(* Logix 5000 project; controller PLC_MCC1300_75F1 vendor 1 type 14 code 166 rev 32.11; software revision 32.04; part 47 of 83 *)
(* tags used below, declared in another part *)
   GP_TrackingFiring : GP_TrackingFiring;
   GP_TrackingFiringForConvoy : GP_TrackingFiringForConvoy;
   M30xTrimWheel : MAC_TrimmingWheels[5];
   M30xTrimWheel_HMR : MAC_TrimmingWheels_HMR[5];
   M30xTrimWheel_HMW : MAC_TrimmingWheels_HMW[5];
   TMP_d : DINT;
   TMP_dIndex : DINT;
   xAlwaysOFF : BOOL;
   Z300_BufferPlate : UDT_LINE_BUFFER_PLATE;
   Z301 : MAC_Zone_ML;
(* MainProgram, continued *)

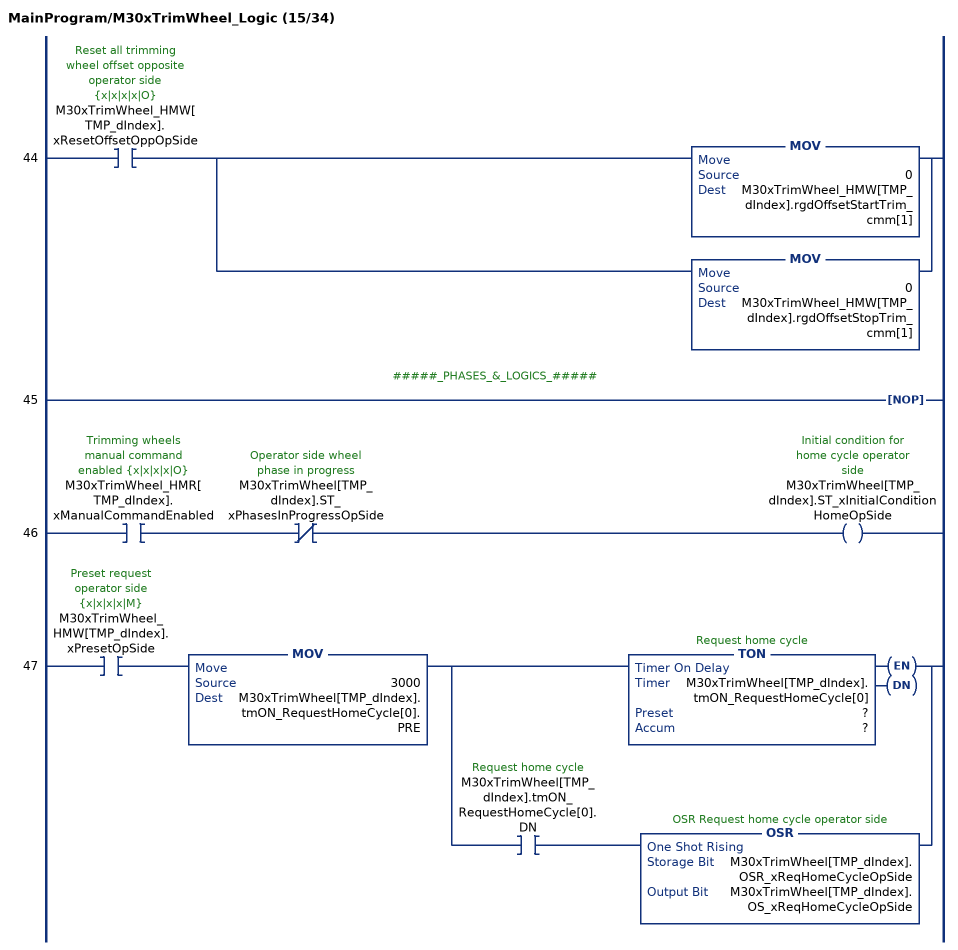
   [picture p701: MainProgram/M30xTrimWheel_Logic rungs 44-47]
   44: XIC(M30xTrimWheel_HMW[TMP_dIndex].xResetOffsetOppOpSide)[MOV(0,M30xTrimWheel_HMW[TMP_dIndex].rgdOffsetStartTrim_cmm[1]) ,MOV(0,M30xTrimWheel_HMW[TMP_dIndex].rgdOffsetStopTrim_cmm[1]) ];
   // #####_PHASES_&_LOGICS_#####
   45: NOP();
   46: XIC(M30xTrimWheel_HMR[TMP_dIndex].xManualCommandEnabled)XIO(M30xTrimWheel[TMP_dIndex].ST_xPhasesInProgressOpSide)OTE(M30xTrimWheel[TMP_dIndex].ST_xInitialConditionHomeOpSide);
   47: XIC(M30xTrimWheel_HMW[TMP_dIndex].xPresetOpSide)MOV(3000,M30xTrimWheel[TMP_dIndex].tmON_RequestHomeCycle[0].PRE)[TON(M30xTrimWheel[TMP_dIndex].tmON_RequestHomeCycle[0],?,?) ,XIC(M30xTrimWheel[TMP_dIndex].tmON_RequestHomeCycle[0].DN) OSR(M30xTrimWheel[TMP_dIndex].OSR_xReqHomeCycleOpSide,M30xTrimWheel[TMP_dIndex].OS_xReqHomeCycleOpSide) ];
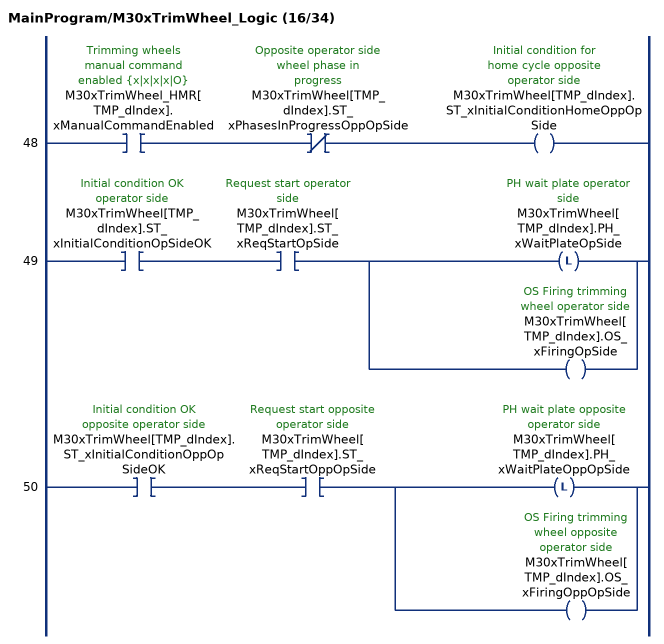
   48: XIC(M30xTrimWheel_HMR[TMP_dIndex].xManualCommandEnabled)XIO(M30xTrimWheel[TMP_dIndex].ST_xPhasesInProgressOppOpSide)OTE(M30xTrimWheel[TMP_dIndex].ST_xInitialConditionHomeOppOpSide);
   49: XIC(M30xTrimWheel[TMP_dIndex].ST_xInitialConditionOpSideOK)XIC(M30xTrimWheel[TMP_dIndex].ST_xReqStartOpSide)[OTL(M30xTrimWheel[TMP_dIndex].PH_xWaitPlateOpSide) ,OTE(M30xTrimWheel[TMP_dIndex].OS_xFiringOpSide) ];
   50: XIC(M30xTrimWheel[TMP_dIndex].ST_xInitialConditionOppOpSideOK)XIC(M30xTrimWheel[TMP_dIndex].ST_xReqStartOppOpSide)[OTL(M30xTrimWheel[TMP_dIndex].PH_xWaitPlateOppOpSide) ,OTE(M30xTrimWheel[TMP_dIndex].OS_xFiringOppOpSide) ];
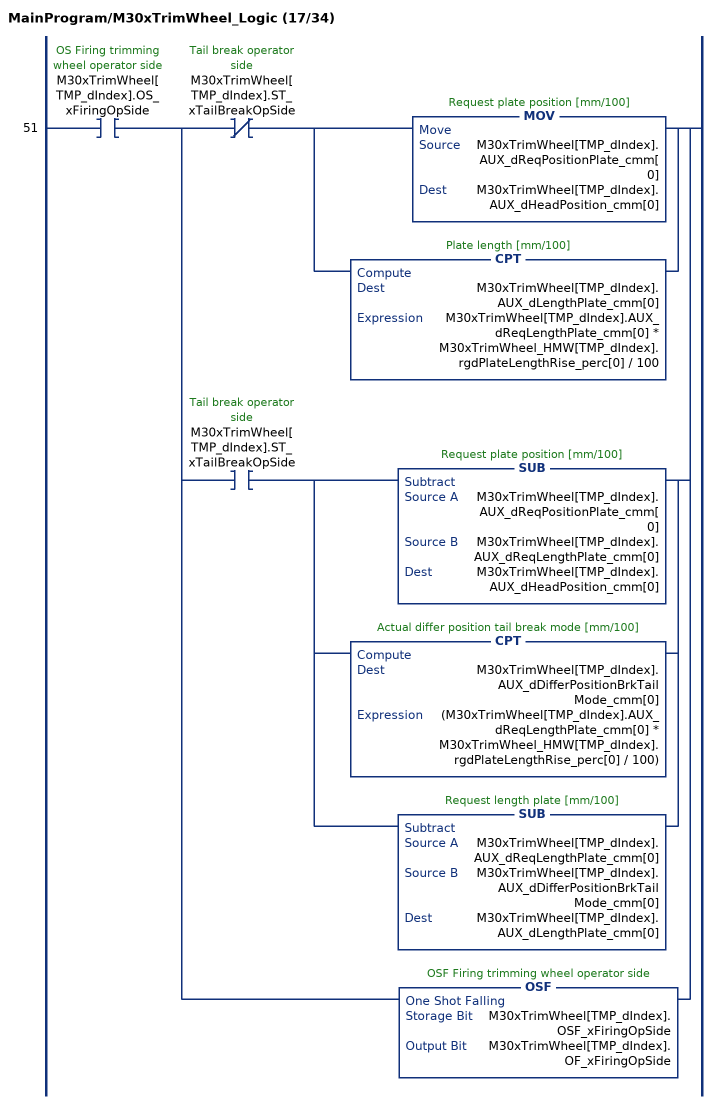
   51: XIC(M30xTrimWheel[TMP_dIndex].OS_xFiringOpSide)[XIO(M30xTrimWheel[TMP_dIndex].ST_xTailBreakOpSide) [MOV(M30xTrimWheel[TMP_dIndex].AUX_dReqPositionPlate_cmm[0],M30xTrimWheel[TMP_dIndex].AUX_dHeadPosition_cmm[0]) ,CPT(M30xTrimWheel[TMP_dIndex].AUX_dLengthPlate_cmm[0],M30xTrimWheel[TMP_dIndex].AUX_dReqLengthPlate_cmm[0] * M30xTrimWheel_HMW[TMP_dIndex].rgdPlateLengthRise_perc[0] / 100) ] ,XIC(M30xTrimWheel[TMP_dIndex].ST_xTailBreakOpSide) [SUB(M30xTrimWheel[TMP_dIndex].AUX_dReqPositionPlate_cmm[0],M30xTrimWheel[TMP_dIndex].AUX_dReqLengthPlate_cmm[0],M30xTrimWheel[TMP_dIndex].AUX_dHeadPosition_cmm[0]) ,CPT(M30xTrimWheel[TMP_dIndex].AUX_dDifferPositionBrkTailMode_cmm[0],(M30xTrimWheel[TMP_dIndex].AUX_dReqLengthPlate_cmm[0] * M30xTrimWheel_HMW[TMP_dIndex].rgdPlateLengthRise_perc[0] / 100)) ,SUB(M30xTrimWheel[TMP_dIndex].AUX_dReqLengthPlate_cmm[0],M30xTrimWheel[TMP_dIndex].AUX_dDifferPositionBrkTailMode_cmm[0],M30xTrimWheel[TMP_dIndex].AUX_dLengthPlate_cmm[0]) ] ,OSF(M30xTrimWheel[TMP_dIndex].OSF_xFiringOpSide,M30xTrimWheel[TMP_dIndex].OF_xFiringOpSide) ];
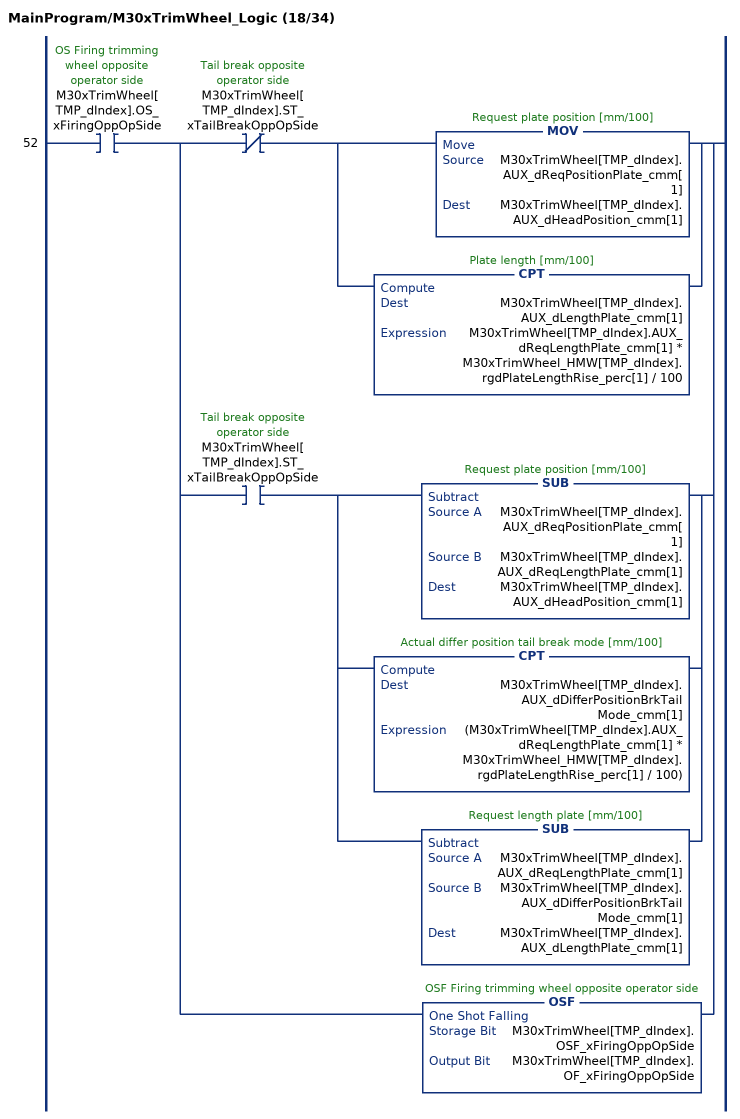
   52: XIC(M30xTrimWheel[TMP_dIndex].OS_xFiringOppOpSide)[XIO(M30xTrimWheel[TMP_dIndex].ST_xTailBreakOppOpSide) [MOV(M30xTrimWheel[TMP_dIndex].AUX_dReqPositionPlate_cmm[1],M30xTrimWheel[TMP_dIndex].AUX_dHeadPosition_cmm[1]) ,CPT(M30xTrimWheel[TMP_dIndex].AUX_dLengthPlate_cmm[1],M30xTrimWheel[TMP_dIndex].AUX_dReqLengthPlate_cmm[1] * M30xTrimWheel_HMW[TMP_dIndex].rgdPlateLengthRise_perc[1] / 100) ] ,XIC(M30xTrimWheel[TMP_dIndex].ST_xTailBreakOppOpSide) [SUB(M30xTrimWheel[TMP_dIndex].AUX_dReqPositionPlate_cmm[1],M30xTrimWheel[TMP_dIndex].AUX_dReqLengthPlate_cmm[1],M30xTrimWheel[TMP_dIndex].AUX_dHeadPosition_cmm[1]) ,CPT(M30xTrimWheel[TMP_dIndex].AUX_dDifferPositionBrkTailMode_cmm[1],(M30xTrimWheel[TMP_dIndex].AUX_dReqLengthPlate_cmm[1] * M30xTrimWheel_HMW[TMP_dIndex].rgdPlateLengthRise_perc[1] / 100)) ,SUB(M30xTrimWheel[TMP_dIndex].AUX_dReqLengthPlate_cmm[1],M30xTrimWheel[TMP_dIndex].AUX_dDifferPositionBrkTailMode_cmm[1],M30xTrimWheel[TMP_dIndex].AUX_dLengthPlate_cmm[1]) ] ,OSF(M30xTrimWheel[TMP_dIndex].OSF_xFiringOppOpSide,M30xTrimWheel[TMP_dIndex].OF_xFiringOppOpSide) ];
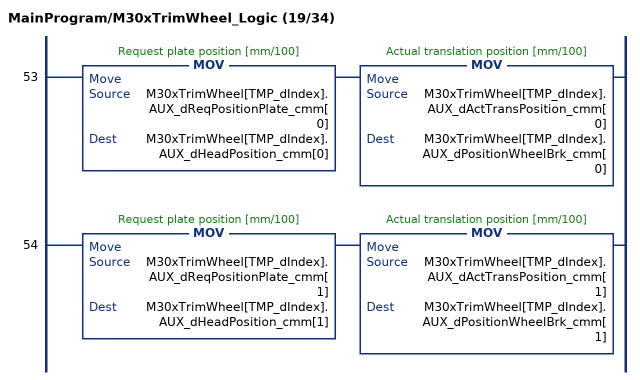
   53: MOV(M30xTrimWheel[TMP_dIndex].AUX_dReqPositionPlate_cmm[0],M30xTrimWheel[TMP_dIndex].AUX_dHeadPosition_cmm[0])MOV(M30xTrimWheel[TMP_dIndex].AUX_dActTransPosition_cmm[0],M30xTrimWheel[TMP_dIndex].AUX_dPositionWheelBrk_cmm[0]);
   54: MOV(M30xTrimWheel[TMP_dIndex].AUX_dReqPositionPlate_cmm[1],M30xTrimWheel[TMP_dIndex].AUX_dHeadPosition_cmm[1])MOV(M30xTrimWheel[TMP_dIndex].AUX_dActTransPosition_cmm[1],M30xTrimWheel[TMP_dIndex].AUX_dPositionWheelBrk_cmm[1]);
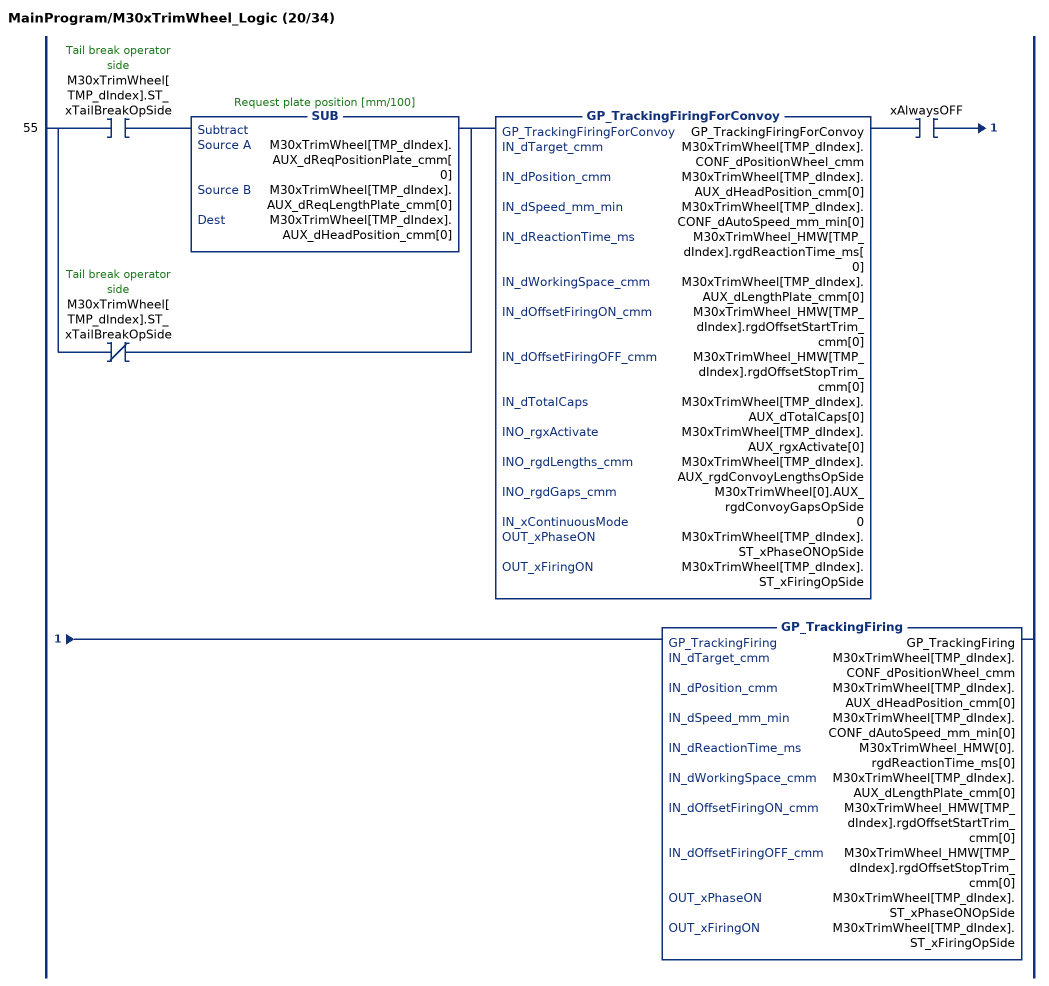
   55: [XIC(M30xTrimWheel[TMP_dIndex].ST_xTailBreakOpSide) SUB(M30xTrimWheel[TMP_dIndex].AUX_dReqPositionPlate_cmm[0],M30xTrimWheel[TMP_dIndex].AUX_dReqLengthPlate_cmm[0],M30xTrimWheel[TMP_dIndex].AUX_dHeadPosition_cmm[0]) ,XIO(M30xTrimWheel[TMP_dIndex].ST_xTailBreakOpSide) ]GP_TrackingFiringForConvoy(GP_TrackingFiringForConvoy,M30xTrimWheel[TMP_dIndex].CONF_dPositionWheel_cmm,M30xTrimWheel[TMP_dIndex].AUX_dHeadPosition_cmm[0],M30xTrimWheel[TMP_dIndex].CONF_dAutoSpeed_mm_min[0],M30xTrimWheel_HMW[TMP_dIndex].rgdReactionTime_ms[0],M30xTrimWheel[TMP_dIndex].AUX_dLengthPlate_cmm[0],M30xTrimWheel_HMW[TMP_dIndex].rgdOffsetStartTrim_cmm[0],M30xTrimWheel_HMW[TMP_dIndex].rgdOffsetStopTrim_cmm[0],M30xTrimWheel[TMP_dIndex].AUX_dTotalCaps[0],M30xTrimWheel[TMP_dIndex].AUX_rgxActivate[0],M30xTrimWheel[TMP_dIndex].AUX_rgdConvoyLengthsOpSide,M30xTrimWheel[0].AUX_rgdConvoyGapsOpSide,0,M30xTrimWheel[TMP_dIndex].ST_xPhaseONOpSide,M30xTrimWheel[TMP_dIndex].ST_xFiringOpSide)XIC(xAlwaysOFF)GP_TrackingFiring(GP_TrackingFiring,M30xTrimWheel[TMP_dIndex].CONF_dPositionWheel_cmm,M30xTrimWheel[TMP_dIndex].AUX_dHeadPosition_cmm[0],M30xTrimWheel[TMP_dIndex].CONF_dAutoSpeed_mm_min[0],M30xTrimWheel_HMW[0].rgdReactionTime_ms[0],M30xTrimWheel[TMP_dIndex].AUX_dLengthPlate_cmm[0],M30xTrimWheel_HMW[TMP_dIndex].rgdOffsetStartTrim_cmm[0],M30xTrimWheel_HMW[TMP_dIndex].rgdOffsetStopTrim_cmm[0],M30xTrimWheel[TMP_dIndex].ST_xPhaseONOpSide,M30xTrimWheel[TMP_dIndex].ST_xFiringOpSide);
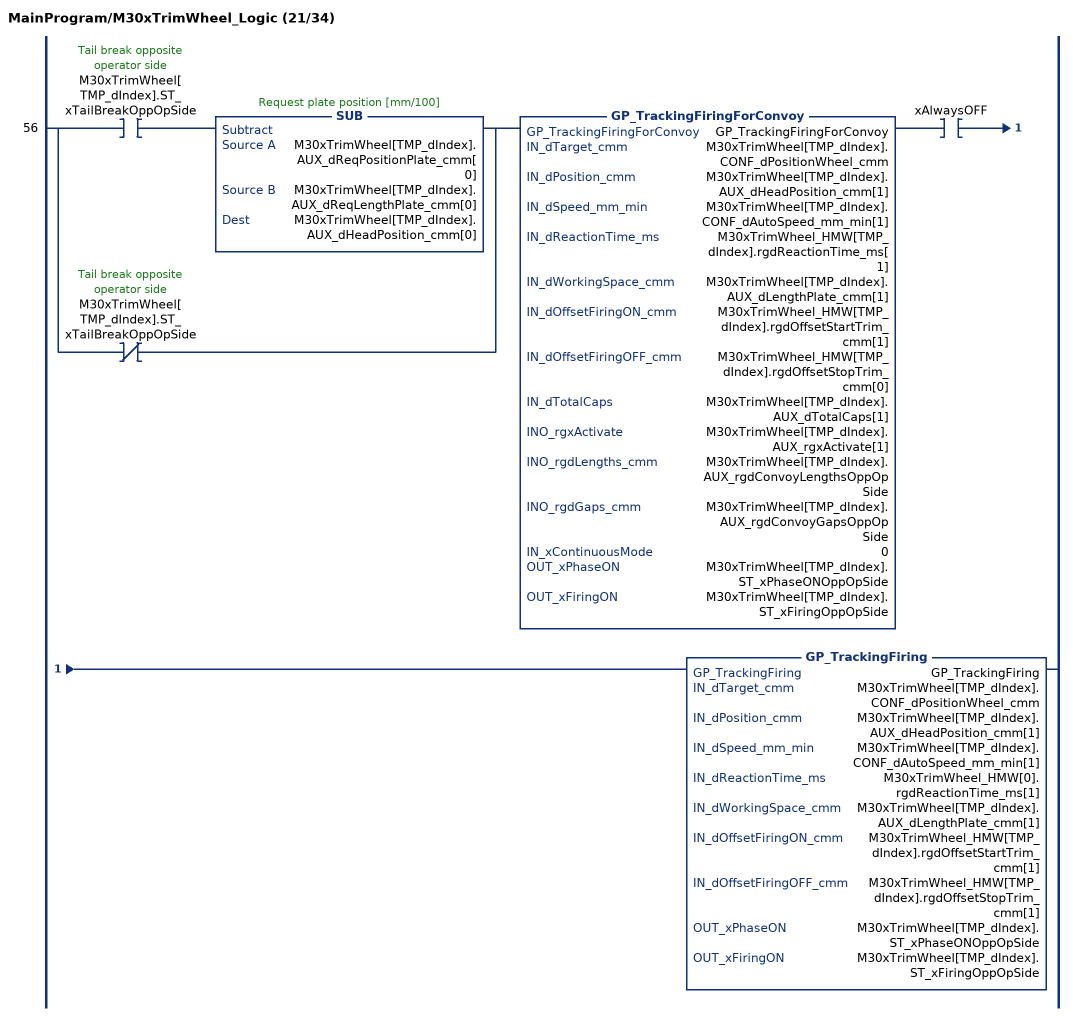
   56: [XIC(M30xTrimWheel[TMP_dIndex].ST_xTailBreakOppOpSide) SUB(M30xTrimWheel[TMP_dIndex].AUX_dReqPositionPlate_cmm[0],M30xTrimWheel[TMP_dIndex].AUX_dReqLengthPlate_cmm[0],M30xTrimWheel[TMP_dIndex].AUX_dHeadPosition_cmm[0]) ,XIO(M30xTrimWheel[TMP_dIndex].ST_xTailBreakOppOpSide) ]GP_TrackingFiringForConvoy(GP_TrackingFiringForConvoy,M30xTrimWheel[TMP_dIndex].CONF_dPositionWheel_cmm,M30xTrimWheel[TMP_dIndex].AUX_dHeadPosition_cmm[1],M30xTrimWheel[TMP_dIndex].CONF_dAutoSpeed_mm_min[1],M30xTrimWheel_HMW[TMP_dIndex].rgdReactionTime_ms[1],M30xTrimWheel[TMP_dIndex].AUX_dLengthPlate_cmm[1],M30xTrimWheel_HMW[TMP_dIndex].rgdOffsetStartTrim_cmm[1],M30xTrimWheel_HMW[TMP_dIndex].rgdOffsetStopTrim_cmm[0],M30xTrimWheel[TMP_dIndex].AUX_dTotalCaps[1],M30xTrimWheel[TMP_dIndex].AUX_rgxActivate[1],M30xTrimWheel[TMP_dIndex].AUX_rgdConvoyLengthsOppOpSide,M30xTrimWheel[TMP_dIndex].AUX_rgdConvoyGapsOppOpSide,0,M30xTrimWheel[TMP_dIndex].ST_xPhaseONOppOpSide,M30xTrimWheel[TMP_dIndex].ST_xFiringOppOpSide)XIC(xAlwaysOFF)GP_TrackingFiring(GP_TrackingFiring,M30xTrimWheel[TMP_dIndex].CONF_dPositionWheel_cmm,M30xTrimWheel[TMP_dIndex].AUX_dHeadPosition_cmm[1],M30xTrimWheel[TMP_dIndex].CONF_dAutoSpeed_mm_min[1],M30xTrimWheel_HMW[0].rgdReactionTime_ms[1],M30xTrimWheel[TMP_dIndex].AUX_dLengthPlate_cmm[1],M30xTrimWheel_HMW[TMP_dIndex].rgdOffsetStartTrim_cmm[1],M30xTrimWheel_HMW[TMP_dIndex].rgdOffsetStopTrim_cmm[1],M30xTrimWheel[TMP_dIndex].ST_xPhaseONOppOpSide,M30xTrimWheel[TMP_dIndex].ST_xFiringOppOpSide);
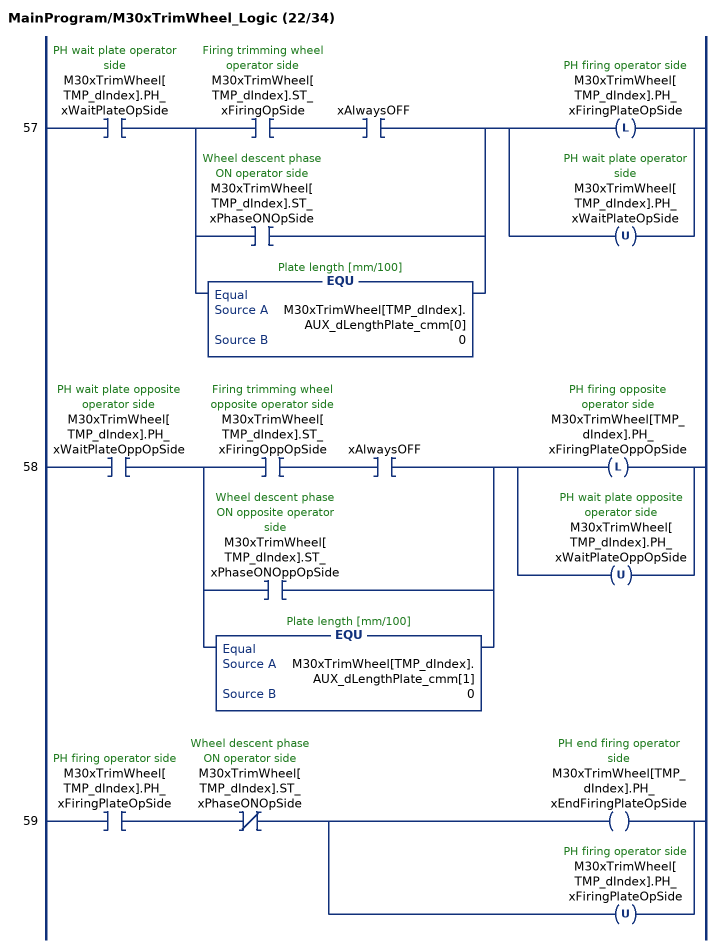
   57: XIC(M30xTrimWheel[TMP_dIndex].PH_xWaitPlateOpSide)[XIC(M30xTrimWheel[TMP_dIndex].ST_xFiringOpSide) XIC(xAlwaysOFF) ,XIC(M30xTrimWheel[TMP_dIndex].ST_xPhaseONOpSide) ,EQU(M30xTrimWheel[TMP_dIndex].AUX_dLengthPlate_cmm[0],0) ][OTL(M30xTrimWheel[TMP_dIndex].PH_xFiringPlateOpSide) ,OTU(M30xTrimWheel[TMP_dIndex].PH_xWaitPlateOpSide) ];
   58: XIC(M30xTrimWheel[TMP_dIndex].PH_xWaitPlateOppOpSide)[XIC(M30xTrimWheel[TMP_dIndex].ST_xFiringOppOpSide) XIC(xAlwaysOFF) ,XIC(M30xTrimWheel[TMP_dIndex].ST_xPhaseONOppOpSide) ,EQU(M30xTrimWheel[TMP_dIndex].AUX_dLengthPlate_cmm[1],0) ][OTL(M30xTrimWheel[TMP_dIndex].PH_xFiringPlateOppOpSide) ,OTU(M30xTrimWheel[TMP_dIndex].PH_xWaitPlateOppOpSide) ];
   59: XIC(M30xTrimWheel[TMP_dIndex].PH_xFiringPlateOpSide)XIO(M30xTrimWheel[TMP_dIndex].ST_xPhaseONOpSide)[OTE(M30xTrimWheel[TMP_dIndex].PH_xEndFiringPlateOpSide) ,OTU(M30xTrimWheel[TMP_dIndex].PH_xFiringPlateOpSide) ];
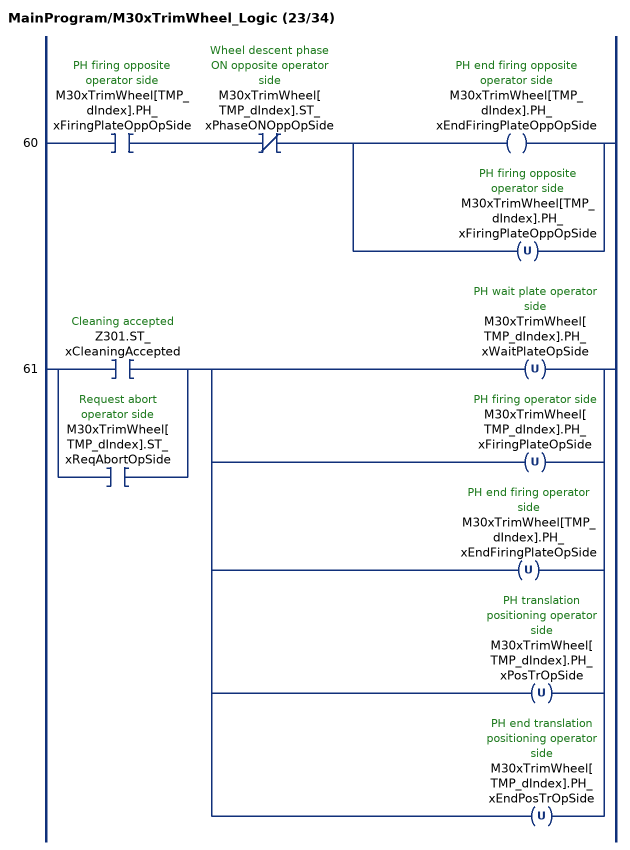
   60: XIC(M30xTrimWheel[TMP_dIndex].PH_xFiringPlateOppOpSide)XIO(M30xTrimWheel[TMP_dIndex].ST_xPhaseONOppOpSide)[OTE(M30xTrimWheel[TMP_dIndex].PH_xEndFiringPlateOppOpSide) ,OTU(M30xTrimWheel[TMP_dIndex].PH_xFiringPlateOppOpSide) ];
   61: [XIC(Z301.ST_xCleaningAccepted) ,XIC(M30xTrimWheel[TMP_dIndex].ST_xReqAbortOpSide) ][OTU(M30xTrimWheel[TMP_dIndex].PH_xWaitPlateOpSide) ,OTU(M30xTrimWheel[TMP_dIndex].PH_xFiringPlateOpSide) ,OTU(M30xTrimWheel[TMP_dIndex].PH_xEndFiringPlateOpSide) ,OTU(M30xTrimWheel[TMP_dIndex].PH_xPosTrOpSide) ,OTU(M30xTrimWheel[TMP_dIndex].PH_xEndPosTrOpSide) ];
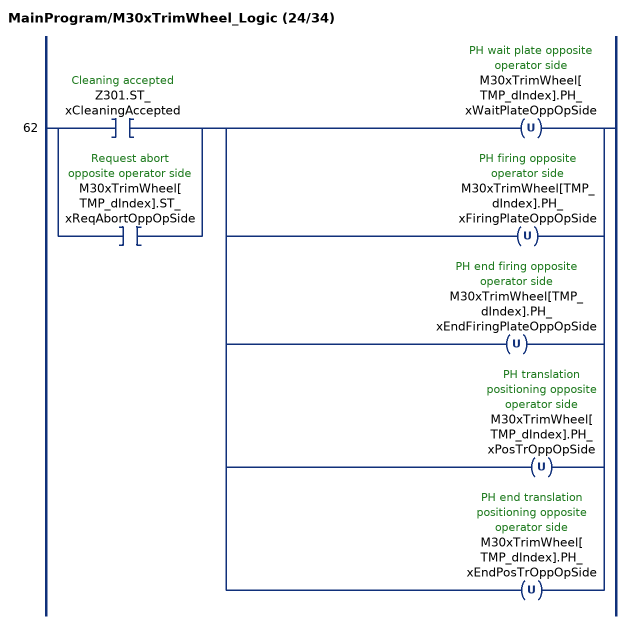
   62: [XIC(Z301.ST_xCleaningAccepted) ,XIC(M30xTrimWheel[TMP_dIndex].ST_xReqAbortOppOpSide) ][OTU(M30xTrimWheel[TMP_dIndex].PH_xWaitPlateOppOpSide) ,OTU(M30xTrimWheel[TMP_dIndex].PH_xFiringPlateOppOpSide) ,OTU(M30xTrimWheel[TMP_dIndex].PH_xEndFiringPlateOppOpSide) ,OTU(M30xTrimWheel[TMP_dIndex].PH_xPosTrOppOpSide) ,OTU(M30xTrimWheel[TMP_dIndex].PH_xEndPosTrOppOpSide) ];
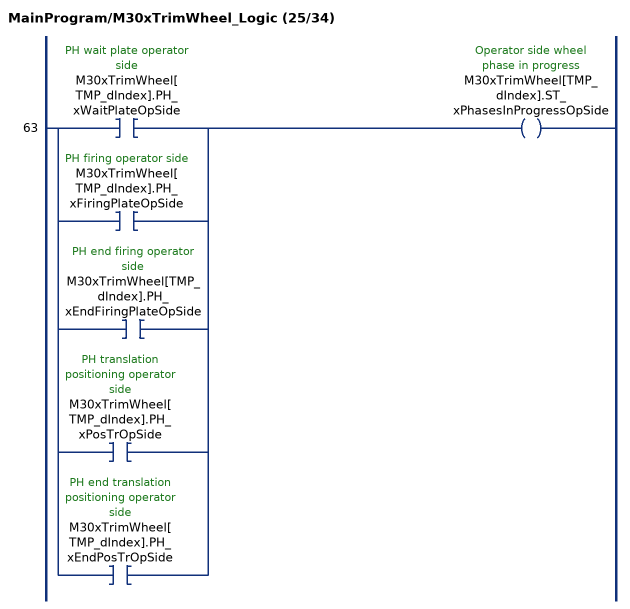
   63: [XIC(M30xTrimWheel[TMP_dIndex].PH_xWaitPlateOpSide) ,XIC(M30xTrimWheel[TMP_dIndex].PH_xFiringPlateOpSide) ,XIC(M30xTrimWheel[TMP_dIndex].PH_xEndFiringPlateOpSide) ,XIC(M30xTrimWheel[TMP_dIndex].PH_xPosTrOpSide) ,XIC(M30xTrimWheel[TMP_dIndex].PH_xEndPosTrOpSide) ]OTE(M30xTrimWheel[TMP_dIndex].ST_xPhasesInProgressOpSide);
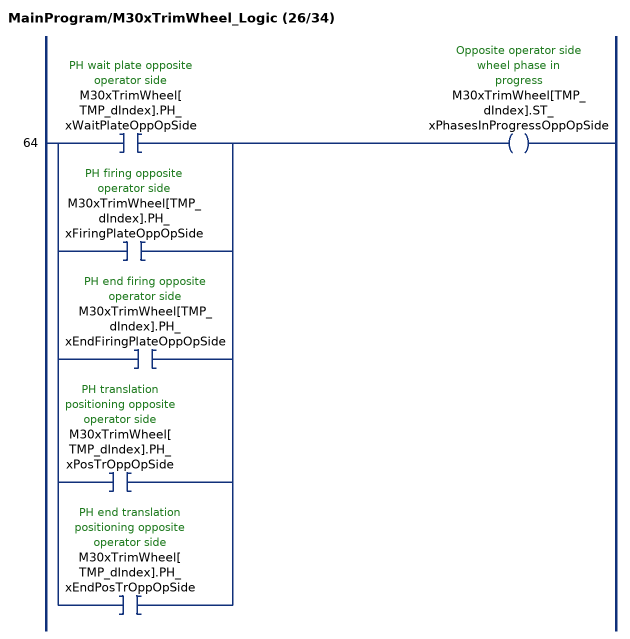
   64: [XIC(M30xTrimWheel[TMP_dIndex].PH_xWaitPlateOppOpSide) ,XIC(M30xTrimWheel[TMP_dIndex].PH_xFiringPlateOppOpSide) ,XIC(M30xTrimWheel[TMP_dIndex].PH_xEndFiringPlateOppOpSide) ,XIC(M30xTrimWheel[TMP_dIndex].PH_xPosTrOppOpSide) ,XIC(M30xTrimWheel[TMP_dIndex].PH_xEndPosTrOppOpSide) ]OTE(M30xTrimWheel[TMP_dIndex].ST_xPhasesInProgressOppOpSide);
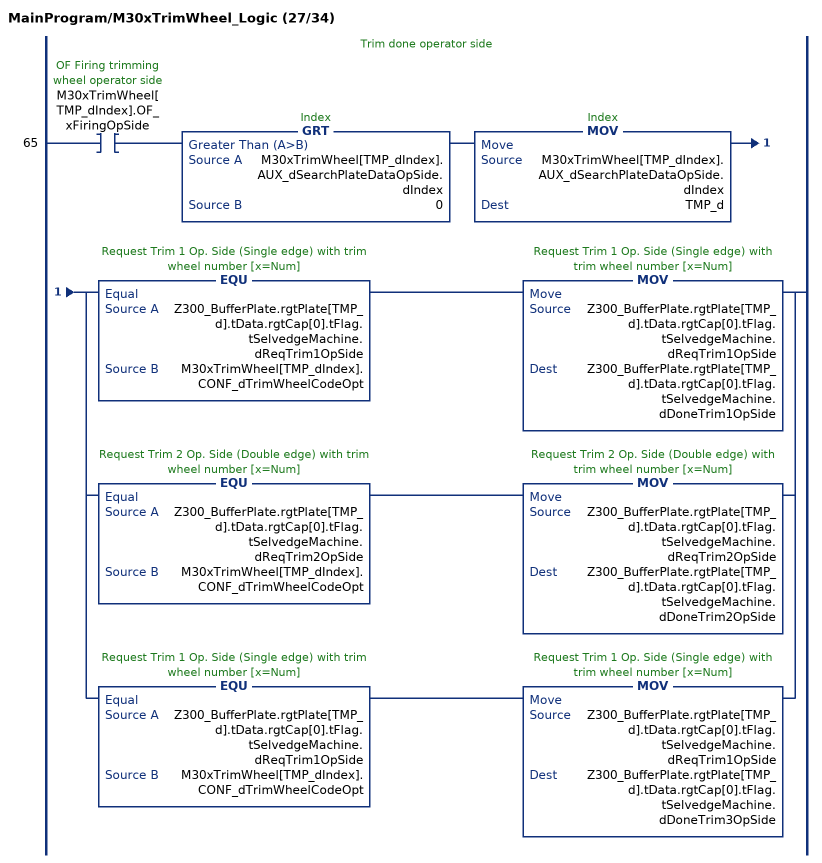
   // Trim done operator side
   65: XIC(M30xTrimWheel[TMP_dIndex].OF_xFiringOpSide)GRT(M30xTrimWheel[TMP_dIndex].AUX_dSearchPlateDataOpSide.dIndex,0)MOV(M30xTrimWheel[TMP_dIndex].AUX_dSearchPlateDataOpSide.dIndex,TMP_d)[EQU(Z300_BufferPlate.rgtPlate[TMP_d].tData.rgtCap[0].tFlag.tSelvedgeMachine.dReqTrim1OpSide,M30xTrimWheel[TMP_dIndex].CONF_dTrimWheelCodeOpt) MOV(Z300_BufferPlate.rgtPlate[TMP_d].tData.rgtCap[0].tFlag.tSelvedgeMachine.dReqTrim1OpSide,Z300_BufferPlate.rgtPlate[TMP_d].tData.rgtCap[0].tFlag.tSelvedgeMachine.dDoneTrim1OpSide) ,EQU(Z300_BufferPlate.rgtPlate[TMP_d].tData.rgtCap[0].tFlag.tSelvedgeMachine.dReqTrim2OpSide,M30xTrimWheel[TMP_dIndex].CONF_dTrimWheelCodeOpt) MOV(Z300_BufferPlate.rgtPlate[TMP_d].tData.rgtCap[0].tFlag.tSelvedgeMachine.dReqTrim2OpSide,Z300_BufferPlate.rgtPlate[TMP_d].tData.rgtCap[0].tFlag.tSelvedgeMachine.dDoneTrim2OpSide) ,EQU(Z300_BufferPlate.rgtPlate[TMP_d].tData.rgtCap[0].tFlag.tSelvedgeMachine.dReqTrim1OpSide,M30xTrimWheel[TMP_dIndex].CONF_dTrimWheelCodeOpt) MOV(Z300_BufferPlate.rgtPlate[TMP_d].tData.rgtCap[0].tFlag.tSelvedgeMachine.dReqTrim1OpSide,Z300_BufferPlate.rgtPlate[TMP_d].tData.rgtCap[0].tFlag.tSelvedgeMachine.dDoneTrim3OpSide) ];
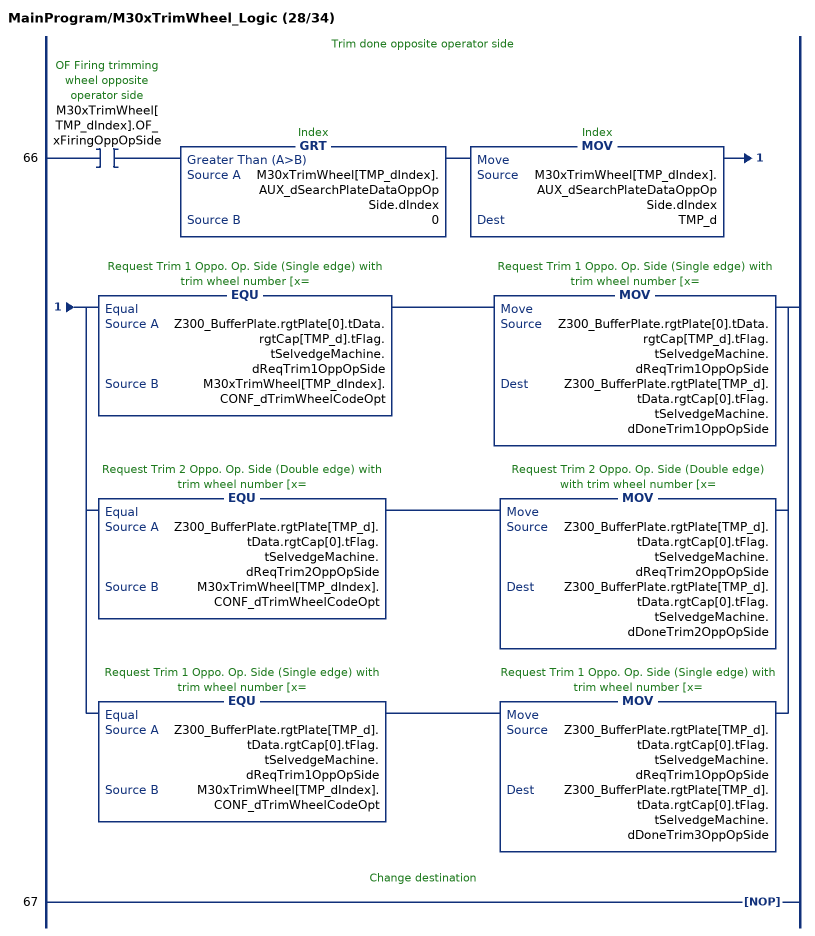
   // Trim done opposite operator side
   66: XIC(M30xTrimWheel[TMP_dIndex].OF_xFiringOppOpSide)GRT(M30xTrimWheel[TMP_dIndex].AUX_dSearchPlateDataOppOpSide.dIndex,0)MOV(M30xTrimWheel[TMP_dIndex].AUX_dSearchPlateDataOppOpSide.dIndex,TMP_d)[EQU(Z300_BufferPlate.rgtPlate[0].tData.rgtCap[TMP_d].tFlag.tSelvedgeMachine.dReqTrim1OppOpSide,M30xTrimWheel[TMP_dIndex].CONF_dTrimWheelCodeOpt) MOV(Z300_BufferPlate.rgtPlate[0].tData.rgtCap[TMP_d].tFlag.tSelvedgeMachine.dReqTrim1OppOpSide,Z300_BufferPlate.rgtPlate[TMP_d].tData.rgtCap[0].tFlag.tSelvedgeMachine.dDoneTrim1OppOpSide) ,EQU(Z300_BufferPlate.rgtPlate[TMP_d].tData.rgtCap[0].tFlag.tSelvedgeMachine.dReqTrim2OppOpSide,M30xTrimWheel[TMP_dIndex].CONF_dTrimWheelCodeOpt) MOV(Z300_BufferPlate.rgtPlate[TMP_d].tData.rgtCap[0].tFlag.tSelvedgeMachine.dReqTrim2OppOpSide,Z300_BufferPlate.rgtPlate[TMP_d].tData.rgtCap[0].tFlag.tSelvedgeMachine.dDoneTrim2OppOpSide) ,EQU(Z300_BufferPlate.rgtPlate[TMP_d].tData.rgtCap[0].tFlag.tSelvedgeMachine.dReqTrim1OppOpSide,M30xTrimWheel[TMP_dIndex].CONF_dTrimWheelCodeOpt) MOV(Z300_BufferPlate.rgtPlate[TMP_d].tData.rgtCap[0].tFlag.tSelvedgeMachine.dReqTrim1OppOpSide,Z300_BufferPlate.rgtPlate[TMP_d].tData.rgtCap[0].tFlag.tSelvedgeMachine.dDoneTrim3OppOpSide) ];
   // Change destination
   67: NOP();
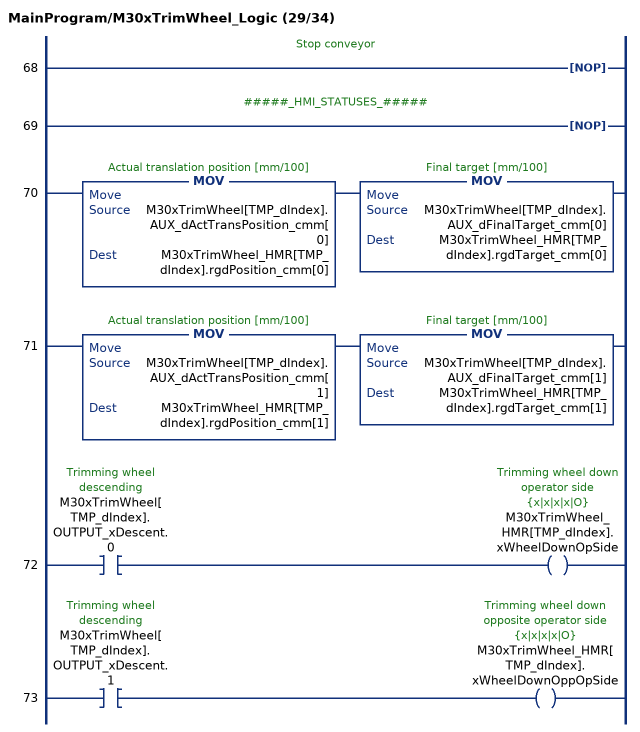
   // Stop conveyor
   68: NOP();
   // #####_HMI_STATUSES_#####
   69: NOP();
   70: MOV(M30xTrimWheel[TMP_dIndex].AUX_dActTransPosition_cmm[0],M30xTrimWheel_HMR[TMP_dIndex].rgdPosition_cmm[0])MOV(M30xTrimWheel[TMP_dIndex].AUX_dFinalTarget_cmm[0],M30xTrimWheel_HMR[TMP_dIndex].rgdTarget_cmm[0]);
   71: MOV(M30xTrimWheel[TMP_dIndex].AUX_dActTransPosition_cmm[1],M30xTrimWheel_HMR[TMP_dIndex].rgdPosition_cmm[1])MOV(M30xTrimWheel[TMP_dIndex].AUX_dFinalTarget_cmm[1],M30xTrimWheel_HMR[TMP_dIndex].rgdTarget_cmm[1]);
   72: XIC(M30xTrimWheel[TMP_dIndex].OUTPUT_xDescent.0)OTE(M30xTrimWheel_HMR[TMP_dIndex].xWheelDownOpSide);
   73: XIC(M30xTrimWheel[TMP_dIndex].OUTPUT_xDescent.1)OTE(M30xTrimWheel_HMR[TMP_dIndex].xWheelDownOppOpSide);
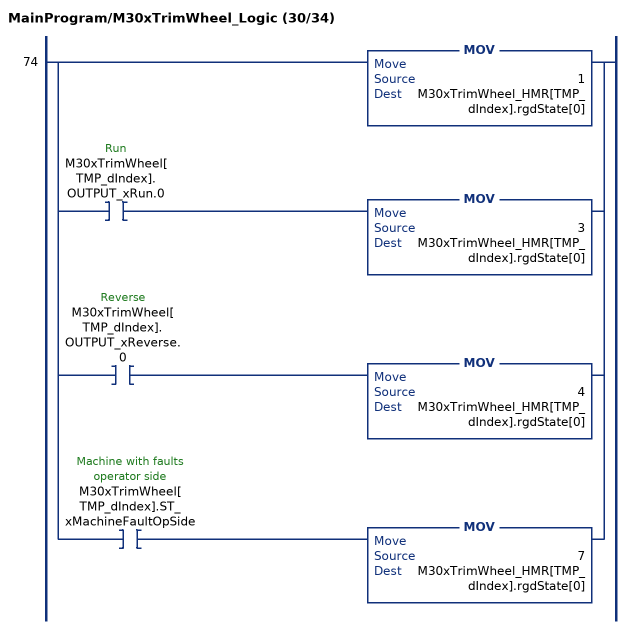
   74: [MOV(1,M30xTrimWheel_HMR[TMP_dIndex].rgdState[0]) ,XIC(M30xTrimWheel[TMP_dIndex].OUTPUT_xRun.0) MOV(3,M30xTrimWheel_HMR[TMP_dIndex].rgdState[0]) ,XIC(M30xTrimWheel[TMP_dIndex].OUTPUT_xReverse.0) MOV(4,M30xTrimWheel_HMR[TMP_dIndex].rgdState[0]) ,XIC(M30xTrimWheel[TMP_dIndex].ST_xMachineFaultOpSide) MOV(7,M30xTrimWheel_HMR[TMP_dIndex].rgdState[0]) ];
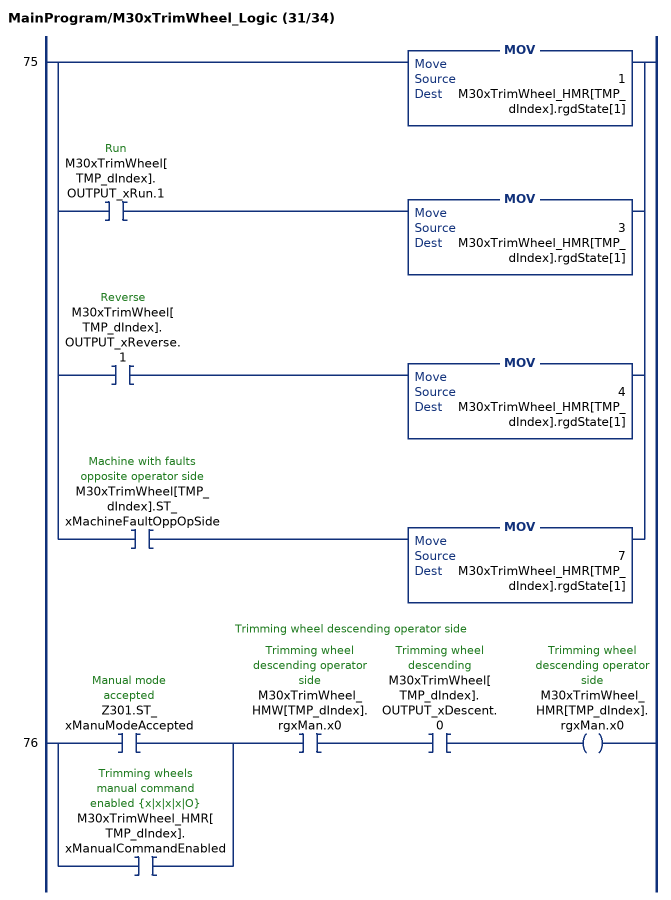
   75: [MOV(1,M30xTrimWheel_HMR[TMP_dIndex].rgdState[1]) ,XIC(M30xTrimWheel[TMP_dIndex].OUTPUT_xRun.1) MOV(3,M30xTrimWheel_HMR[TMP_dIndex].rgdState[1]) ,XIC(M30xTrimWheel[TMP_dIndex].OUTPUT_xReverse.1) MOV(4,M30xTrimWheel_HMR[TMP_dIndex].rgdState[1]) ,XIC(M30xTrimWheel[TMP_dIndex].ST_xMachineFaultOppOpSide) MOV(7,M30xTrimWheel_HMR[TMP_dIndex].rgdState[1]) ];
   // Trimming wheel descending operator side
   76: [XIC(Z301.ST_xManuModeAccepted) ,XIC(M30xTrimWheel_HMR[TMP_dIndex].xManualCommandEnabled) ]XIC(M30xTrimWheel_HMW[TMP_dIndex].rgxMan.x0)XIC(M30xTrimWheel[TMP_dIndex].OUTPUT_xDescent.0)OTE(M30xTrimWheel_HMR[TMP_dIndex].rgxMan.x0);
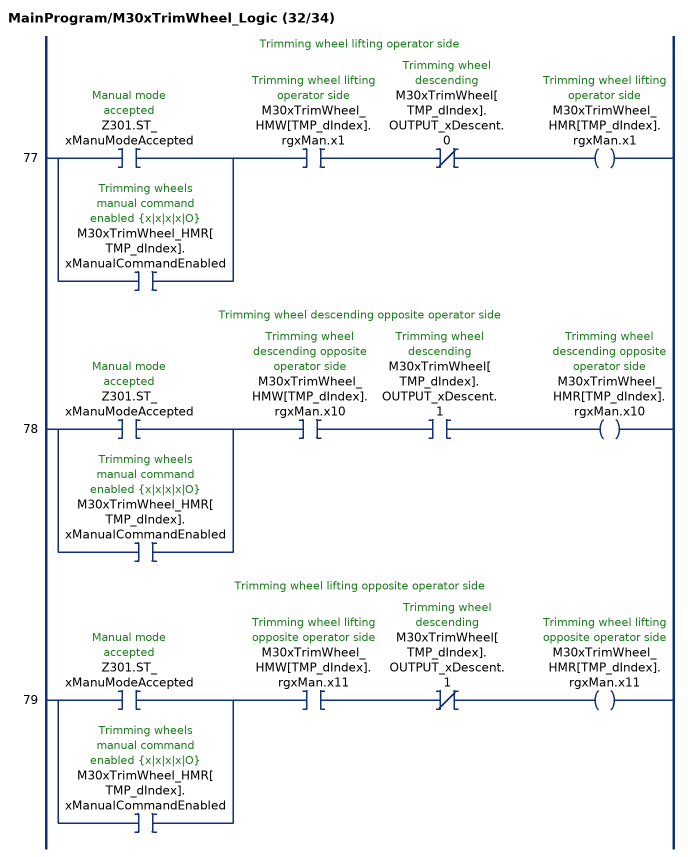
   // Trimming wheel lifting operator side
   77: [XIC(Z301.ST_xManuModeAccepted) ,XIC(M30xTrimWheel_HMR[TMP_dIndex].xManualCommandEnabled) ]XIC(M30xTrimWheel_HMW[TMP_dIndex].rgxMan.x1)XIO(M30xTrimWheel[TMP_dIndex].OUTPUT_xDescent.0)OTE(M30xTrimWheel_HMR[TMP_dIndex].rgxMan.x1);
   // Trimming wheel descending opposite operator side
   78: [XIC(Z301.ST_xManuModeAccepted) ,XIC(M30xTrimWheel_HMR[TMP_dIndex].xManualCommandEnabled) ]XIC(M30xTrimWheel_HMW[TMP_dIndex].rgxMan.x10)XIC(M30xTrimWheel[TMP_dIndex].OUTPUT_xDescent.1)OTE(M30xTrimWheel_HMR[TMP_dIndex].rgxMan.x10);
   // Trimming wheel lifting opposite operator side
   79: [XIC(Z301.ST_xManuModeAccepted) ,XIC(M30xTrimWheel_HMR[TMP_dIndex].xManualCommandEnabled) ]XIC(M30xTrimWheel_HMW[TMP_dIndex].rgxMan.x11)XIO(M30xTrimWheel[TMP_dIndex].OUTPUT_xDescent.1)OTE(M30xTrimWheel_HMR[TMP_dIndex].rgxMan.x11);
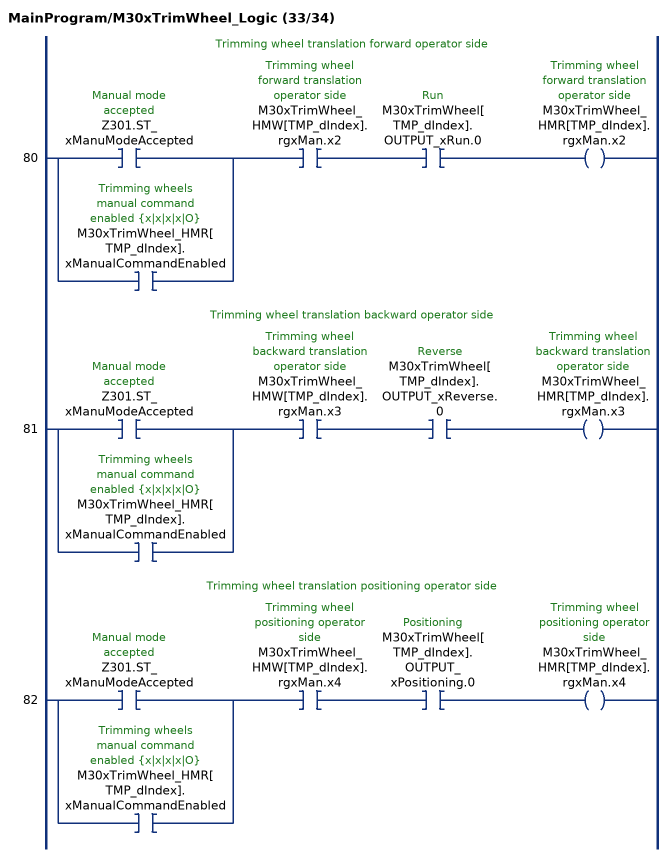
   // Trimming wheel translation forward operator side
   80: [XIC(Z301.ST_xManuModeAccepted) ,XIC(M30xTrimWheel_HMR[TMP_dIndex].xManualCommandEnabled) ]XIC(M30xTrimWheel_HMW[TMP_dIndex].rgxMan.x2)XIC(M30xTrimWheel[TMP_dIndex].OUTPUT_xRun.0)OTE(M30xTrimWheel_HMR[TMP_dIndex].rgxMan.x2);
   // Trimming wheel translation backward operator side
   81: [XIC(Z301.ST_xManuModeAccepted) ,XIC(M30xTrimWheel_HMR[TMP_dIndex].xManualCommandEnabled) ]XIC(M30xTrimWheel_HMW[TMP_dIndex].rgxMan.x3)XIC(M30xTrimWheel[TMP_dIndex].OUTPUT_xReverse.0)OTE(M30xTrimWheel_HMR[TMP_dIndex].rgxMan.x3);
   // Trimming wheel translation positioning operator side
   82: [XIC(Z301.ST_xManuModeAccepted) ,XIC(M30xTrimWheel_HMR[TMP_dIndex].xManualCommandEnabled) ]XIC(M30xTrimWheel_HMW[TMP_dIndex].rgxMan.x4)XIC(M30xTrimWheel[TMP_dIndex].OUTPUT_xPositioning.0)OTE(M30xTrimWheel_HMR[TMP_dIndex].rgxMan.x4);
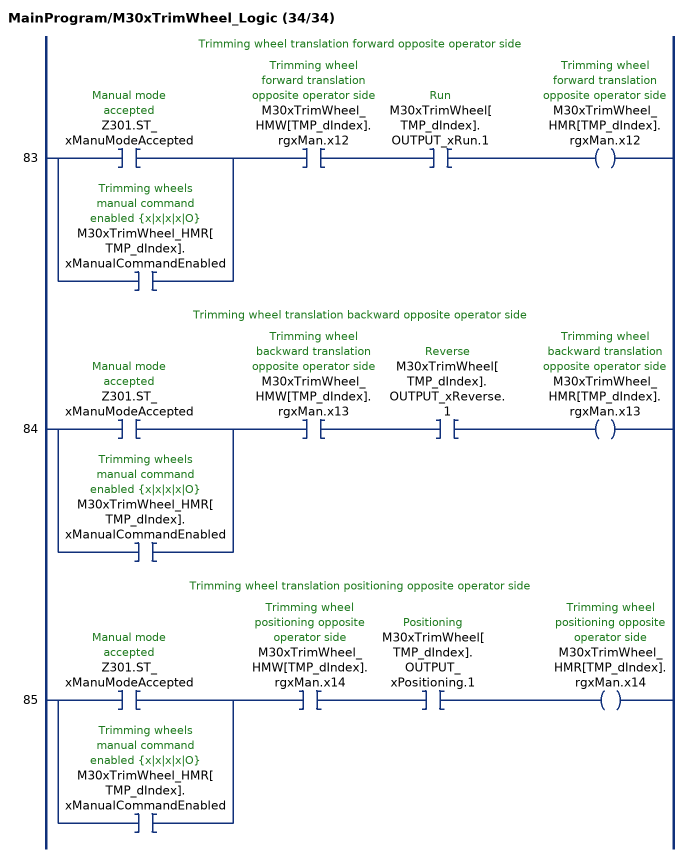
   // Trimming wheel translation forward opposite operator side
   83: [XIC(Z301.ST_xManuModeAccepted) ,XIC(M30xTrimWheel_HMR[TMP_dIndex].xManualCommandEnabled) ]XIC(M30xTrimWheel_HMW[TMP_dIndex].rgxMan.x12)XIC(M30xTrimWheel[TMP_dIndex].OUTPUT_xRun.1)OTE(M30xTrimWheel_HMR[TMP_dIndex].rgxMan.x12);
   // Trimming wheel translation backward opposite operator side
   84: [XIC(Z301.ST_xManuModeAccepted) ,XIC(M30xTrimWheel_HMR[TMP_dIndex].xManualCommandEnabled) ]XIC(M30xTrimWheel_HMW[TMP_dIndex].rgxMan.x13)XIC(M30xTrimWheel[TMP_dIndex].OUTPUT_xReverse.1)OTE(M30xTrimWheel_HMR[TMP_dIndex].rgxMan.x13);
   // Trimming wheel translation positioning opposite operator side
   85: [XIC(Z301.ST_xManuModeAccepted) ,XIC(M30xTrimWheel_HMR[TMP_dIndex].xManualCommandEnabled) ]XIC(M30xTrimWheel_HMW[TMP_dIndex].rgxMan.x14)XIC(M30xTrimWheel[TMP_dIndex].OUTPUT_xPositioning.1)OTE(M30xTrimWheel_HMR[TMP_dIndex].rgxMan.x14);
END_ROUTINE
